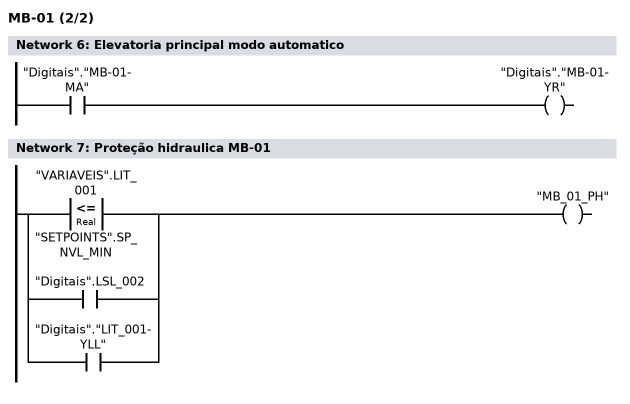
   RUNG wire#powerrail
      Contact( "Digitais"."MB-01-MA" )
      Coil( "Digitais"."MB-01-YR" )
   END_RUNG
   // the same network as SCL:
   "Digitais"."MB-01-YR" := "Digitais"."MB-01-MA";
END_REGION

REGION Network 7: Proteção hidraulica MB-01
   RUNG wire#powerrail
      { S7_Templates := "SrcType := Real" } LE_Contact(in1 := "VARIAVEIS".LIT_001, in2 := "SETPOINTS".SP_NVL_MIN)
      wire#w1
      Coil( "MB_01_PH" )
   END_RUNG
   RUNG wire#powerrail
      Contact( "Digitais".LSL_002 )
   END_RUNG wire#w1
   RUNG wire#powerrail
      Contact( "Digitais"."LIT_001-YLL" )
   END_RUNG wire#w1
   // the same network as SCL:
   "MB_01_PH" := ("VARIAVEIS".LIT_001 <= "SETPOINTS".SP_NVL_MIN) OR "Digitais".LSL_002 OR "Digitais"."LIT_001-YLL";
END_REGION
END_FUNCTION

FUNCTION "MB-02" : Void   // FC23, LAD
TITLE = Lógica de acionamento do motor
{ S7_Optimized_Access := 'FALSE' }
VERSION : 0.1
   VAR_TEMP
      IM : Bool;   // Intertravamento manual = 0
      IA : Bool;   // Intertravamento automáticol = 0
      HABM : Bool;   // Habilita funcionamento manual = 1
      HABA : Bool;   // Habilita funcionamento automático = 1
      CLM : Bool;   // Comando liga motor
      PROT : Bool;   // Proteção do motor acionada
   END_VAR
BEGIN

REGION Network 1: Intertravamento maual/automático
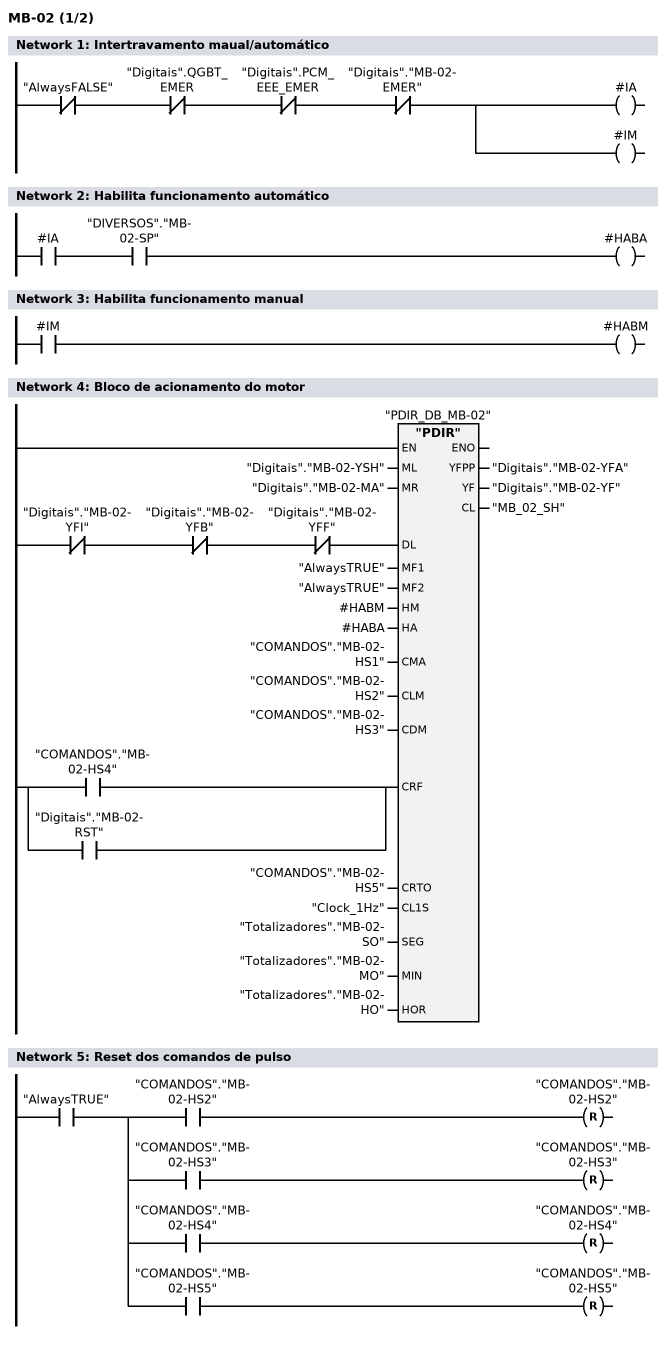
   RUNG wire#powerrail
      I_Contact( "AlwaysFALSE" )
      I_Contact( "Digitais".QGBT_EMER )
      I_Contact( "Digitais".PCM_EEE_EMER )
      I_Contact( "Digitais"."MB-02-EMER" )
      wire#w1
      Coil( #IA )
   END_RUNG
   RUNG wire#w1
      Coil( #IM )
   END_RUNG
   // the same network as SCL:
   #IA := NOT "AlwaysFALSE" AND NOT "Digitais".QGBT_EMER AND NOT "Digitais".PCM_EEE_EMER AND NOT "Digitais"."MB-02-EMER";
   #IM := #IA;
END_REGION

REGION Network 2: Habilita funcionamento automático
   RUNG wire#powerrail
      Contact( #IA )
      Contact( "DIVERSOS"."MB-02-SP" )
      Coil( #HABA )
   END_RUNG
   // the same network as SCL:
   #HABA := #IA AND "DIVERSOS"."MB-02-SP";
END_REGION

REGION Network 3: Habilita funcionamento manual
   RUNG wire#powerrail
      Contact( #IM )
      Coil( #HABM )
   END_RUNG
   // the same network as SCL:
   #HABM := #IM;
END_REGION

REGION Network 4: Bloco de acionamento do motor
   RUNG wire#powerrail
      "PDIR_DB_MB-02"(DL := wire#w1, CRF := wire#w2, ML := "Digitais"."MB-02-YSH", MR := "Digitais"."MB-02-MA", MF1 := "AlwaysTRUE", MF2 := "AlwaysTRUE", HM := #HABM, HA := #HABA, CMA := "COMANDOS"."MB-02-HS1", CLM := "COMANDOS"."MB-02-HS2", CDM := "COMANDOS"."MB-02-HS3", CRTO := "COMANDOS"."MB-02-HS5", CL1S := "Clock_1Hz", SEG := "Totalizadores"."MB-02-SO", MIN := "Totalizadores"."MB-02-MO", HOR := "Totalizadores"."MB-02-HO", YFPP => "Digitais"."MB-02-YFA", YF => "Digitais"."MB-02-YF", CL => "MB_02_SH")
   END_RUNG
   RUNG wire#powerrail
      I_Contact( "Digitais"."MB-02-YFI" )
      I_Contact( "Digitais"."MB-02-YFB" )
      I_Contact( "Digitais"."MB-02-YFF" )
   END_RUNG wire#w1
   RUNG wire#powerrail
      Contact( "COMANDOS"."MB-02-HS4" )
   END_RUNG wire#w2
   RUNG wire#powerrail
      Contact( "Digitais"."MB-02-RST" )
   END_RUNG wire#w2
   // the same network as SCL:
   "PDIR_DB_MB-02"(ML := "Digitais"."MB-02-YSH",   // "PDIR"
                   MR := "Digitais"."MB-02-MA",
                   DL := NOT "Digitais"."MB-02-YFI" AND NOT "Digitais"."MB-02-YFB" AND NOT "Digitais"."MB-02-YFF",
                   MF1 := "AlwaysTRUE",
                   MF2 := "AlwaysTRUE",
                   HM := #HABM,
                   HA := #HABA,
                   CMA := "COMANDOS"."MB-02-HS1",
                   CLM := "COMANDOS"."MB-02-HS2",
                   CDM := "COMANDOS"."MB-02-HS3",
                   CRF := "COMANDOS"."MB-02-HS4" OR "Digitais"."MB-02-RST",
                   CRTO := "COMANDOS"."MB-02-HS5",
                   CL1S := "Clock_1Hz",
                   SEG := "Totalizadores"."MB-02-SO",
                   MIN := "Totalizadores"."MB-02-MO",
                   HOR := "Totalizadores"."MB-02-HO",
                   YFPP => "Digitais"."MB-02-YFA",
                   YF => "Digitais"."MB-02-YF",
                   CL => "MB_02_SH");
END_REGION

REGION Network 5: Reset dos comandos de pulso
   RUNG wire#powerrail
      Contact( "AlwaysTRUE" )
      wire#w1
      Contact( "COMANDOS"."MB-02-HS2" )
      R_Coil( "COMANDOS"."MB-02-HS2" )
   END_RUNG
   RUNG wire#w1
      Contact( "COMANDOS"."MB-02-HS3" )
      R_Coil( "COMANDOS"."MB-02-HS3" )
   END_RUNG
   RUNG wire#w1
      Contact( "COMANDOS"."MB-02-HS4" )
      R_Coil( "COMANDOS"."MB-02-HS4" )
   END_RUNG
   RUNG wire#w1
      Contact( "COMANDOS"."MB-02-HS5" )
      R_Coil( "COMANDOS"."MB-02-HS5" )
   END_RUNG
   // the same network as SCL:
   IF "AlwaysTRUE" AND "COMANDOS"."MB-02-HS2" THEN "COMANDOS"."MB-02-HS2" := FALSE; END_IF;
   IF "AlwaysTRUE" AND "COMANDOS"."MB-02-HS3" THEN "COMANDOS"."MB-02-HS3" := FALSE; END_IF;
   IF "AlwaysTRUE" AND "COMANDOS"."MB-02-HS4" THEN "COMANDOS"."MB-02-HS4" := FALSE; END_IF;
   IF "AlwaysTRUE" AND "COMANDOS"."MB-02-HS5" THEN "COMANDOS"."MB-02-HS5" := FALSE; END_IF;
END_REGION

REGION Network 6: Elevatoria principal modo automatico
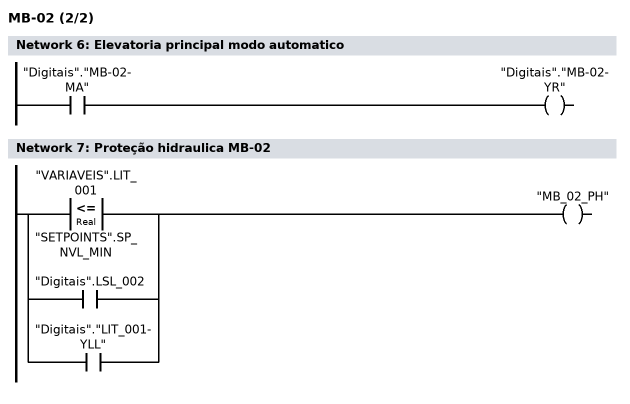
   RUNG wire#powerrail
      Contact( "Digitais"."MB-02-MA" )
      Coil( "Digitais"."MB-02-YR" )
   END_RUNG
   // the same network as SCL:
   "Digitais"."MB-02-YR" := "Digitais"."MB-02-MA";
END_REGION

REGION Network 7: Proteção hidraulica MB-02
   RUNG wire#powerrail
      { S7_Templates := "SrcType := Real" } LE_Contact(in1 := "VARIAVEIS".LIT_001, in2 := "SETPOINTS".SP_NVL_MIN)
      wire#w1
      Coil( "MB_02_PH" )
   END_RUNG
   RUNG wire#powerrail
      Contact( "Digitais".LSL_002 )
   END_RUNG wire#w1
   RUNG wire#powerrail
      Contact( "Digitais"."LIT_001-YLL" )
   END_RUNG wire#w1
   // the same network as SCL:
   "MB_02_PH" := ("VARIAVEIS".LIT_001 <= "SETPOINTS".SP_NVL_MIN) OR "Digitais".LSL_002 OR "Digitais"."LIT_001-YLL";
END_REGION
END_FUNCTION

FUNCTION "MB-03" : Void   // FC24, LAD
TITLE = Lógica de acionamento do motor
{ S7_Optimized_Access := 'FALSE' }
VERSION : 0.1
   VAR_TEMP
      IM : Bool;   // Intertravamento manual = 0
      IA : Bool;   // Intertravamento automáticol = 0
      HABM : Bool;   // Habilita funcionamento manual = 1
      HABA : Bool;   // Habilita funcionamento automático = 1
      CLM : Bool;   // Comando liga motor
      PROT : Bool;   // Proteção do motor acionada
   END_VAR
BEGIN

REGION Network 1: Intertravamento maual/automático
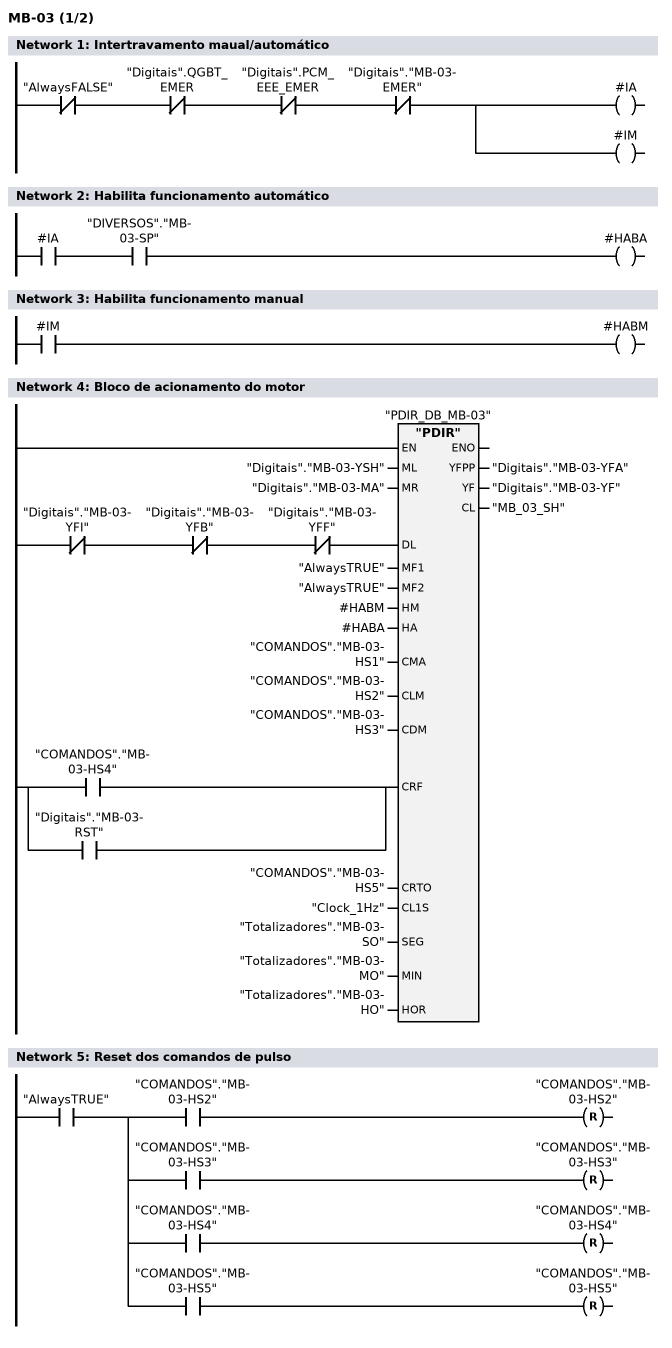
   RUNG wire#powerrail
      I_Contact( "AlwaysFALSE" )
      I_Contact( "Digitais".QGBT_EMER )
      I_Contact( "Digitais".PCM_EEE_EMER )
      I_Contact( "Digitais"."MB-03-EMER" )
      wire#w1
      Coil( #IA )
   END_RUNG
   RUNG wire#w1
      Coil( #IM )
   END_RUNG
   // the same network as SCL:
   #IA := NOT "AlwaysFALSE" AND NOT "Digitais".QGBT_EMER AND NOT "Digitais".PCM_EEE_EMER AND NOT "Digitais"."MB-03-EMER";
   #IM := #IA;
END_REGION

REGION Network 2: Habilita funcionamento automático
   RUNG wire#powerrail
      Contact( #IA )
      Contact( "DIVERSOS"."MB-03-SP" )
      Coil( #HABA )
   END_RUNG
   // the same network as SCL:
   #HABA := #IA AND "DIVERSOS"."MB-03-SP";
END_REGION

REGION Network 3: Habilita funcionamento manual
   RUNG wire#powerrail
      Contact( #IM )
      Coil( #HABM )
   END_RUNG
   // the same network as SCL:
   #HABM := #IM;
END_REGION

REGION Network 4: Bloco de acionamento do motor
   RUNG wire#powerrail
      "PDIR_DB_MB-03"(DL := wire#w1, CRF := wire#w2, ML := "Digitais"."MB-03-YSH", MR := "Digitais"."MB-03-MA", MF1 := "AlwaysTRUE", MF2 := "AlwaysTRUE", HM := #HABM, HA := #HABA, CMA := "COMANDOS"."MB-03-HS1", CLM := "COMANDOS"."MB-03-HS2", CDM := "COMANDOS"."MB-03-HS3", CRTO := "COMANDOS"."MB-03-HS5", CL1S := "Clock_1Hz", SEG := "Totalizadores"."MB-03-SO", MIN := "Totalizadores"."MB-03-MO", HOR := "Totalizadores"."MB-03-HO", YFPP => "Digitais"."MB-03-YFA", YF => "Digitais"."MB-03-YF", CL => "MB_03_SH")
   END_RUNG
   RUNG wire#powerrail
      I_Contact( "Digitais"."MB-03-YFI" )
      I_Contact( "Digitais"."MB-03-YFB" )
      I_Contact( "Digitais"."MB-03-YFF" )
   END_RUNG wire#w1
   RUNG wire#powerrail
      Contact( "COMANDOS"."MB-03-HS4" )
   END_RUNG wire#w2
   RUNG wire#powerrail
      Contact( "Digitais"."MB-03-RST" )
   END_RUNG wire#w2
   // the same network as SCL:
   "PDIR_DB_MB-03"(ML := "Digitais"."MB-03-YSH",   // "PDIR"
                   MR := "Digitais"."MB-03-MA",
                   DL := NOT "Digitais"."MB-03-YFI" AND NOT "Digitais"."MB-03-YFB" AND NOT "Digitais"."MB-03-YFF",
                   MF1 := "AlwaysTRUE",
                   MF2 := "AlwaysTRUE",
                   HM := #HABM,
                   HA := #HABA,
                   CMA := "COMANDOS"."MB-03-HS1",
                   CLM := "COMANDOS"."MB-03-HS2",
                   CDM := "COMANDOS"."MB-03-HS3",
                   CRF := "COMANDOS"."MB-03-HS4" OR "Digitais"."MB-03-RST",
                   CRTO := "COMANDOS"."MB-03-HS5",
                   CL1S := "Clock_1Hz",
                   SEG := "Totalizadores"."MB-03-SO",
                   MIN := "Totalizadores"."MB-03-MO",
                   HOR := "Totalizadores"."MB-03-HO",
                   YFPP => "Digitais"."MB-03-YFA",
                   YF => "Digitais"."MB-03-YF",
                   CL => "MB_03_SH");
END_REGION

REGION Network 5: Reset dos comandos de pulso
   RUNG wire#powerrail
      Contact( "AlwaysTRUE" )
      wire#w1
      Contact( "COMANDOS"."MB-03-HS2" )
      R_Coil( "COMANDOS"."MB-03-HS2" )
   END_RUNG
   RUNG wire#w1
      Contact( "COMANDOS"."MB-03-HS3" )
      R_Coil( "COMANDOS"."MB-03-HS3" )
   END_RUNG
   RUNG wire#w1
      Contact( "COMANDOS"."MB-03-HS4" )
      R_Coil( "COMANDOS"."MB-03-HS4" )
   END_RUNG
   RUNG wire#w1
      Contact( "COMANDOS"."MB-03-HS5" )
      R_Coil( "COMANDOS"."MB-03-HS5" )
   END_RUNG
   // the same network as SCL:
   IF "AlwaysTRUE" AND "COMANDOS"."MB-03-HS2" THEN "COMANDOS"."MB-03-HS2" := FALSE; END_IF;
   IF "AlwaysTRUE" AND "COMANDOS"."MB-03-HS3" THEN "COMANDOS"."MB-03-HS3" := FALSE; END_IF;
   IF "AlwaysTRUE" AND "COMANDOS"."MB-03-HS4" THEN "COMANDOS"."MB-03-HS4" := FALSE; END_IF;
   IF "AlwaysTRUE" AND "COMANDOS"."MB-03-HS5" THEN "COMANDOS"."MB-03-HS5" := FALSE; END_IF;
END_REGION

REGION Network 6: Elevatoria principal modo automatico
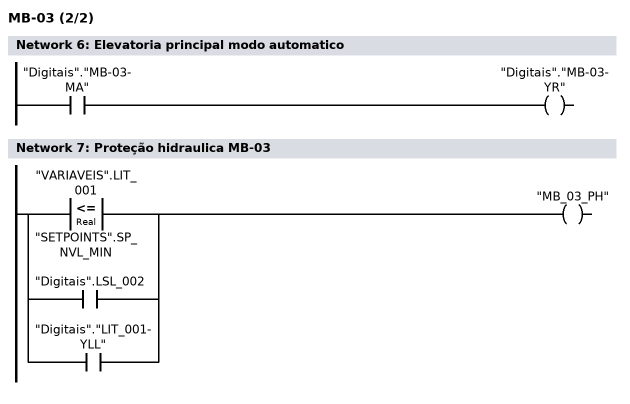
   RUNG wire#powerrail
      Contact( "Digitais"."MB-03-MA" )
      Coil( "Digitais"."MB-03-YR" )
   END_RUNG
   // the same network as SCL:
   "Digitais"."MB-03-YR" := "Digitais"."MB-03-MA";
END_REGION

REGION Network 7: Proteção hidraulica MB-03
   RUNG wire#powerrail
      { S7_Templates := "SrcType := Real" } LE_Contact(in1 := "VARIAVEIS".LIT_001, in2 := "SETPOINTS".SP_NVL_MIN)
      wire#w1
      Coil( "MB_03_PH" )
   END_RUNG
   RUNG wire#powerrail
      Contact( "Digitais".LSL_002 )
   END_RUNG wire#w1
   RUNG wire#powerrail
      Contact( "Digitais"."LIT_001-YLL" )
   END_RUNG wire#w1
   // the same network as SCL:
   "MB_03_PH" := ("VARIAVEIS".LIT_001 <= "SETPOINTS".SP_NVL_MIN) OR "Digitais".LSL_002 OR "Digitais"."LIT_001-YLL";
END_REGION
END_FUNCTION

FUNCTION "MB-04" : Void   // FC25, LAD
TITLE = Lógica de acionamento do motor
{ S7_Optimized_Access := 'FALSE' }
VERSION : 0.1
   VAR_TEMP
      IM : Bool;   // Intertravamento manual = 0
      IA : Bool;   // Intertravamento automáticol = 0
      HABM : Bool;   // Habilita funcionamento manual = 1
      HABA : Bool;   // Habilita funcionamento automático = 1
      CLM : Bool;   // Comando liga motor
      PROT : Bool;   // Proteção do motor acionada
   END_VAR
BEGIN

REGION Network 1: Intertravamento maual/automático
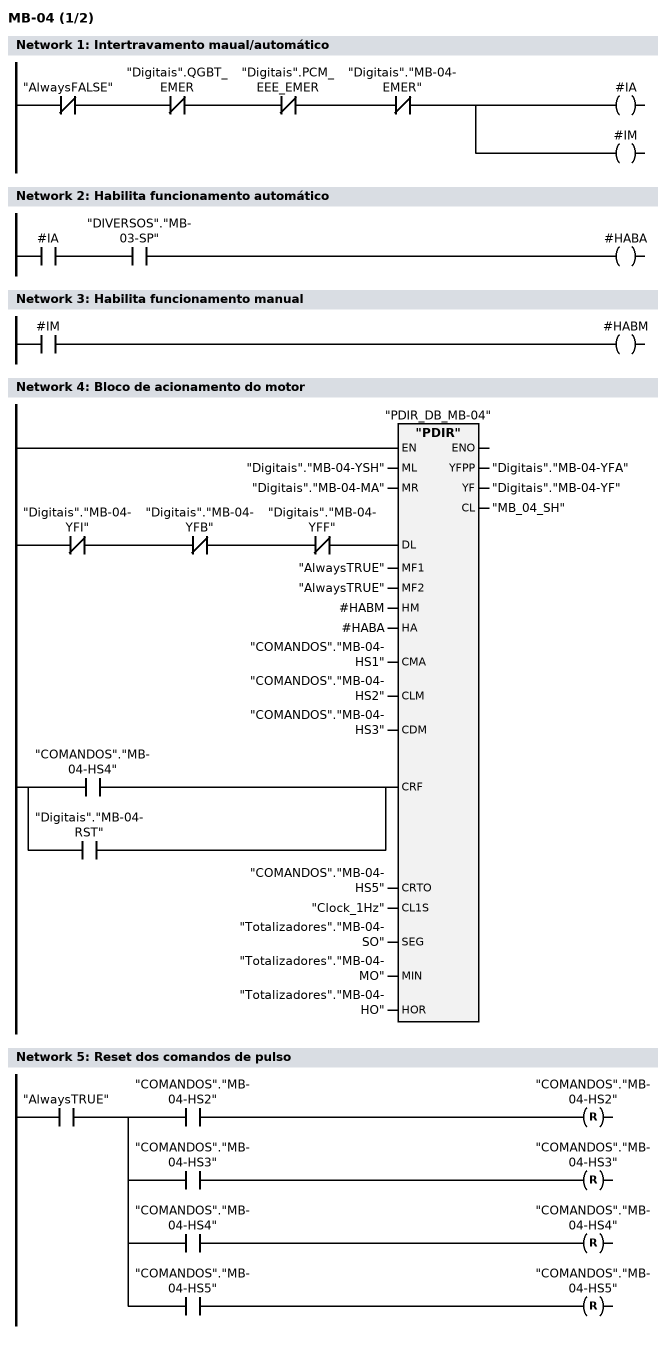
   RUNG wire#powerrail
      I_Contact( "AlwaysFALSE" )
      I_Contact( "Digitais".QGBT_EMER )
      I_Contact( "Digitais".PCM_EEE_EMER )
      I_Contact( "Digitais"."MB-04-EMER" )
      wire#w1
      Coil( #IA )
   END_RUNG
   RUNG wire#w1
      Coil( #IM )
   END_RUNG
   // the same network as SCL:
   #IA := NOT "AlwaysFALSE" AND NOT "Digitais".QGBT_EMER AND NOT "Digitais".PCM_EEE_EMER AND NOT "Digitais"."MB-04-EMER";
   #IM := #IA;
END_REGION

REGION Network 2: Habilita funcionamento automático
   RUNG wire#powerrail
      Contact( #IA )
      Contact( "DIVERSOS"."MB-03-SP" )
      Coil( #HABA )
   END_RUNG
   // the same network as SCL:
   #HABA := #IA AND "DIVERSOS"."MB-03-SP";
END_REGION

REGION Network 3: Habilita funcionamento manual
   RUNG wire#powerrail
      Contact( #IM )
      Coil( #HABM )
   END_RUNG
   // the same network as SCL:
   #HABM := #IM;
END_REGION

REGION Network 4: Bloco de acionamento do motor
   RUNG wire#powerrail
      "PDIR_DB_MB-04"(DL := wire#w1, CRF := wire#w2, ML := "Digitais"."MB-04-YSH", MR := "Digitais"."MB-04-MA", MF1 := "AlwaysTRUE", MF2 := "AlwaysTRUE", HM := #HABM, HA := #HABA, CMA := "COMANDOS"."MB-04-HS1", CLM := "COMANDOS"."MB-04-HS2", CDM := "COMANDOS"."MB-04-HS3", CRTO := "COMANDOS"."MB-04-HS5", CL1S := "Clock_1Hz", SEG := "Totalizadores"."MB-04-SO", MIN := "Totalizadores"."MB-04-MO", HOR := "Totalizadores"."MB-04-HO", YFPP => "Digitais"."MB-04-YFA", YF => "Digitais"."MB-04-YF", CL => "MB_04_SH")
   END_RUNG
   RUNG wire#powerrail
      I_Contact( "Digitais"."MB-04-YFI" )
      I_Contact( "Digitais"."MB-04-YFB" )
      I_Contact( "Digitais"."MB-04-YFF" )
   END_RUNG wire#w1
   RUNG wire#powerrail
      Contact( "COMANDOS"."MB-04-HS4" )
   END_RUNG wire#w2
   RUNG wire#powerrail
      Contact( "Digitais"."MB-04-RST" )
   END_RUNG wire#w2
   // the same network as SCL:
   "PDIR_DB_MB-04"(ML := "Digitais"."MB-04-YSH",   // "PDIR"
                   MR := "Digitais"."MB-04-MA",
                   DL := NOT "Digitais"."MB-04-YFI" AND NOT "Digitais"."MB-04-YFB" AND NOT "Digitais"."MB-04-YFF",
                   MF1 := "AlwaysTRUE",
                   MF2 := "AlwaysTRUE",
                   HM := #HABM,
                   HA := #HABA,
                   CMA := "COMANDOS"."MB-04-HS1",
                   CLM := "COMANDOS"."MB-04-HS2",
                   CDM := "COMANDOS"."MB-04-HS3",
                   CRF := "COMANDOS"."MB-04-HS4" OR "Digitais"."MB-04-RST",
                   CRTO := "COMANDOS"."MB-04-HS5",
                   CL1S := "Clock_1Hz",
                   SEG := "Totalizadores"."MB-04-SO",
                   MIN := "Totalizadores"."MB-04-MO",
                   HOR := "Totalizadores"."MB-04-HO",
                   YFPP => "Digitais"."MB-04-YFA",
                   YF => "Digitais"."MB-04-YF",
                   CL => "MB_04_SH");
END_REGION

REGION Network 5: Reset dos comandos de pulso
   RUNG wire#powerrail
      Contact( "AlwaysTRUE" )
      wire#w1
      Contact( "COMANDOS"."MB-04-HS2" )
      R_Coil( "COMANDOS"."MB-04-HS2" )
   END_RUNG
   RUNG wire#w1
      Contact( "COMANDOS"."MB-04-HS3" )
      R_Coil( "COMANDOS"."MB-04-HS3" )
   END_RUNG
   RUNG wire#w1
      Contact( "COMANDOS"."MB-04-HS4" )
      R_Coil( "COMANDOS"."MB-04-HS4" )
   END_RUNG
   RUNG wire#w1
      Contact( "COMANDOS"."MB-04-HS5" )
      R_Coil( "COMANDOS"."MB-04-HS5" )
   END_RUNG
   // the same network as SCL:
   IF "AlwaysTRUE" AND "COMANDOS"."MB-04-HS2" THEN "COMANDOS"."MB-04-HS2" := FALSE; END_IF;
   IF "AlwaysTRUE" AND "COMANDOS"."MB-04-HS3" THEN "COMANDOS"."MB-04-HS3" := FALSE; END_IF;
   IF "AlwaysTRUE" AND "COMANDOS"."MB-04-HS4" THEN "COMANDOS"."MB-04-HS4" := FALSE; END_IF;
   IF "AlwaysTRUE" AND "COMANDOS"."MB-04-HS5" THEN "COMANDOS"."MB-04-HS5" := FALSE; END_IF;
END_REGION

REGION Network 6: Elevatoria principal modo automatico
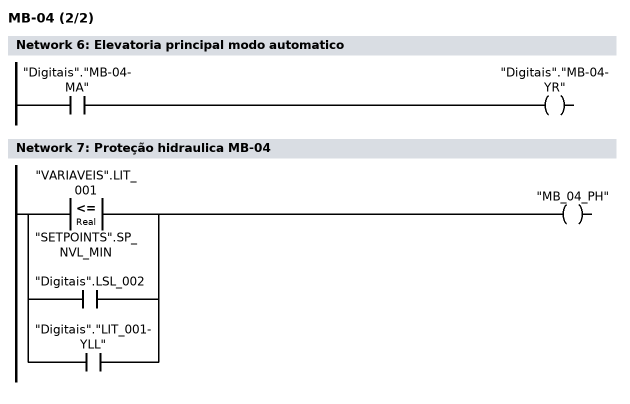
   RUNG wire#powerrail
      Contact( "Digitais"."MB-04-MA" )
      Coil( "Digitais"."MB-04-YR" )
   END_RUNG
   // the same network as SCL:
   "Digitais"."MB-04-YR" := "Digitais"."MB-04-MA";
END_REGION

REGION Network 7: Proteção hidraulica MB-04
   RUNG wire#powerrail
      { S7_Templates := "SrcType := Real" } LE_Contact(in1 := "VARIAVEIS".LIT_001, in2 := "SETPOINTS".SP_NVL_MIN)
      wire#w1
      Coil( "MB_04_PH" )
   END_RUNG
   RUNG wire#powerrail
      Contact( "Digitais".LSL_002 )
   END_RUNG wire#w1
   RUNG wire#powerrail
      Contact( "Digitais"."LIT_001-YLL" )
   END_RUNG wire#w1
   // the same network as SCL:
   "MB_04_PH" := ("VARIAVEIS".LIT_001 <= "SETPOINTS".SP_NVL_MIN) OR "Digitais".LSL_002 OR "Digitais"."LIT_001-YLL";
END_REGION
END_FUNCTION

ORGANIZATION_BLOCK "Main"   // OB1, LAD, ProgramCycle
TITLE = "Main Program Sweep (Cycle)"
{ S7_Optimized_Access := 'TRUE' }
VERSION : 0.1
   VAR_INPUT
      Initial_Call : Bool;   // Initial call of this OB
      Remanence : Bool;   // =True, if remanent data are available
   END_VAR
BEGIN

REGION Network 1: PULSO 1 SEGUNDO
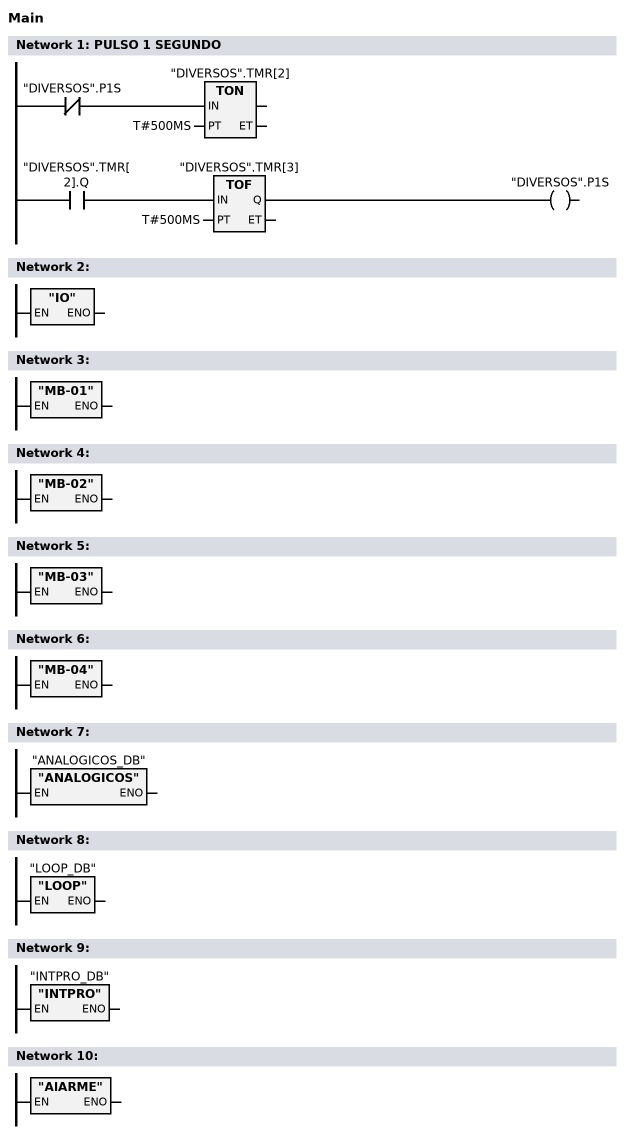
   "DIVERSOS".TMR[2].TON(IN := NOT "DIVERSOS".P1S, PT := T#500MS);
   "DIVERSOS".TMR[3].TOF(IN := "DIVERSOS".TMR[2].Q, PT := T#500MS);
   "DIVERSOS".P1S := "DIVERSOS".TMR[3].Q;
END_REGION

REGION Network 2
   RUNG wire#powerrail
      "IO"()
   END_RUNG
   // the same network as SCL:
   "IO"();
END_REGION

REGION Network 3
   RUNG wire#powerrail
      "MB-01"()
   END_RUNG
   // the same network as SCL:
   "MB-01"();
END_REGION

REGION Network 4
   RUNG wire#powerrail
      "MB-02"()
   END_RUNG
   // the same network as SCL:
   "MB-02"();
END_REGION

REGION Network 5
   RUNG wire#powerrail
      "MB-03"()
   END_RUNG
   // the same network as SCL:
   "MB-03"();
END_REGION

REGION Network 6
   RUNG wire#powerrail
      "MB-04"()
   END_RUNG
   // the same network as SCL:
   "MB-04"();
END_REGION

REGION Network 7
   RUNG wire#powerrail
      "ANALOGICOS_DB"()
   END_RUNG
   // the same network as SCL:
   "ANALOGICOS_DB"();   // "ANALOGICOS"
END_REGION

REGION Network 8
   RUNG wire#powerrail
      "LOOP_DB"()
   END_RUNG
   // the same network as SCL:
   "LOOP_DB"();   // "LOOP"
END_REGION

REGION Network 9
   RUNG wire#powerrail
      "INTPRO_DB"()
   END_RUNG
   // the same network as SCL:
   "INTPRO_DB"();   // "INTPRO"
END_REGION

REGION Network 10
   RUNG wire#powerrail
      "AlARME"()
   END_RUNG
   // the same network as SCL:
   "AlARME"();
END_REGION
END_ORGANIZATION_BLOCK

ORGANIZATION_BLOCK "CYC_INT5"   // OB35, LAD, CyclicInterrupt
TITLE = CONTROLE DE PID
{ S7_Optimized_Access := 'FALSE' }
VERSION : 0.1
   VAR_TEMP
      OB35_EV_CLASS : Byte;
      OB35_STRT_INF : Byte;
      OB35_PRIORITY : Byte;
      OB35_OB_NUMBR : Byte;
      OB35_RESERVED_1 : Byte;
      OB35_RESERVED_2 : Byte;
      OB35_PHASE_OFFSET : Word;
      OB35_RESERVED_3 : Int;
      OB35_EXC_FREQ : Int;
      OB35_DATE_TIME : Date_And_Time;
      "SPM-EEEB" : Real;   // Setpoint manual PID tanque de aeração 1
      EEEB_IT : Time;   // Ajuste integral do PID
      EEEB_DT : Time;   // Ajuste derivativo do PID
      EEEB_AUX : Real;   // Setpoint manual PID - auxiliar
      EEEB_P : Real;   // Setpoint manual PID - auxiliar
   END_VAR
   VAR_TEMP   // added for the SCL form of the ladder/FBD networks
      _w1 : Bool;
      _w2 : Bool;
      _w3 : Bool;
      _w4 : Bool;
   END_VAR
BEGIN

REGION Network 1 (STL): CONVERSÃO DOS SETPOINTS PARA TEMPO PID EEEB


   //CONVERSÃO DOS SETPOINTS DE TEMPO PID EEEB
         L     "PID"."PID-EEEB-I";
         L     1000.0;
         *R;
         RND;
         T     #EEEB_IT;

         L     "PID"."PID-EEEB-D";
         L     1000.0;
         *R;
         RND;
         T     #EEEB_DT;

         L     "PID"."PID-EEEB-P";
         L     -1.0;
         *R;
         T     #EEEB_P;
END_REGION

REGION Network 2: PID TANQUE DE AERAÇÃO 1
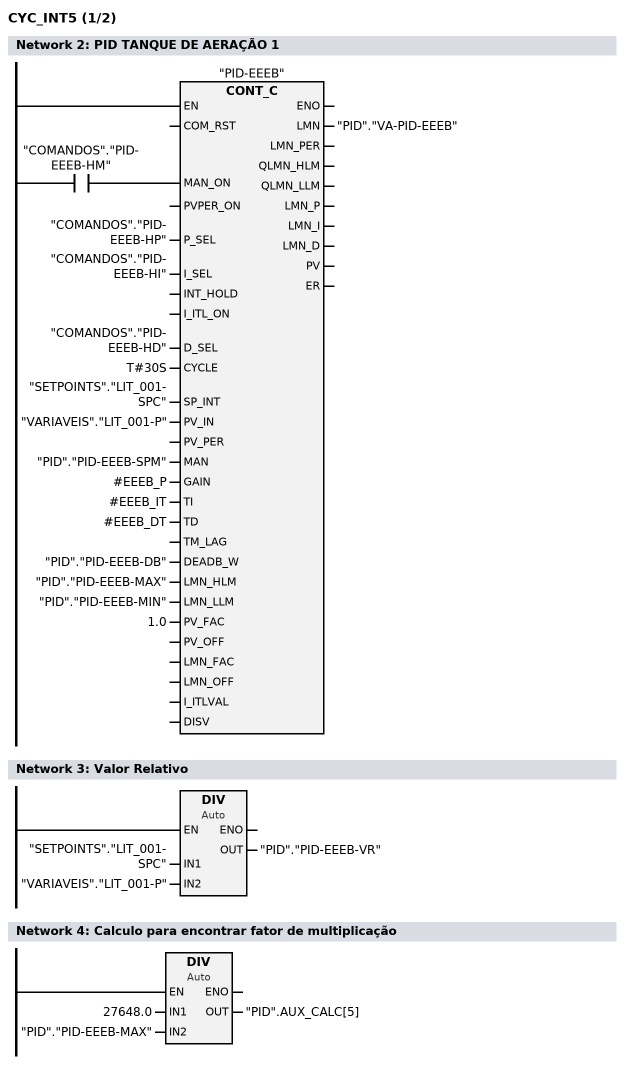
   "PID-EEEB"(MAN_ON := "COMANDOS"."PID-EEEB-HM",   // CONT_C
              P_SEL := "COMANDOS"."PID-EEEB-HP",
              I_SEL := "COMANDOS"."PID-EEEB-HI",
              D_SEL := "COMANDOS"."PID-EEEB-HD",
              CYCLE := T#30S,
              SP_INT := "SETPOINTS"."LIT_001-SPC",
              PV_IN := "VARIAVEIS"."LIT_001-P",
              MAN := "PID"."PID-EEEB-SPM",
              GAIN := #EEEB_P,
              TI := #EEEB_IT,
              TD := #EEEB_DT,
              DEADB_W := "PID"."PID-EEEB-DB",
              LMN_HLM := "PID"."PID-EEEB-MAX",
              LMN_LLM := "PID"."PID-EEEB-MIN",
              PV_FAC := 1.0,
              LMN => "PID"."VA-PID-EEEB");
END_REGION

REGION Network 3: Valor Relativo
   RUNG wire#powerrail
      Div(in1 := "SETPOINTS"."LIT_001-SPC", in2 := "VARIAVEIS"."LIT_001-P", out => "PID"."PID-EEEB-VR")
   END_RUNG
   // the same network as SCL:
   "PID"."PID-EEEB-VR" := "SETPOINTS"."LIT_001-SPC" / "VARIAVEIS"."LIT_001-P";
END_REGION

REGION Network 4: Calculo para encontrar fator de multiplicação
   RUNG wire#powerrail
      Div(in1 := 27648.0, in2 := "PID"."PID-EEEB-MAX", out => "PID".AUX_CALC[5])
   END_RUNG
   // the same network as SCL:
   "PID".AUX_CALC[5] := 27648.0 / "PID"."PID-EEEB-MAX";
END_REGION

REGION Network 5: Movimenta saida PID para entrada analógica inversor
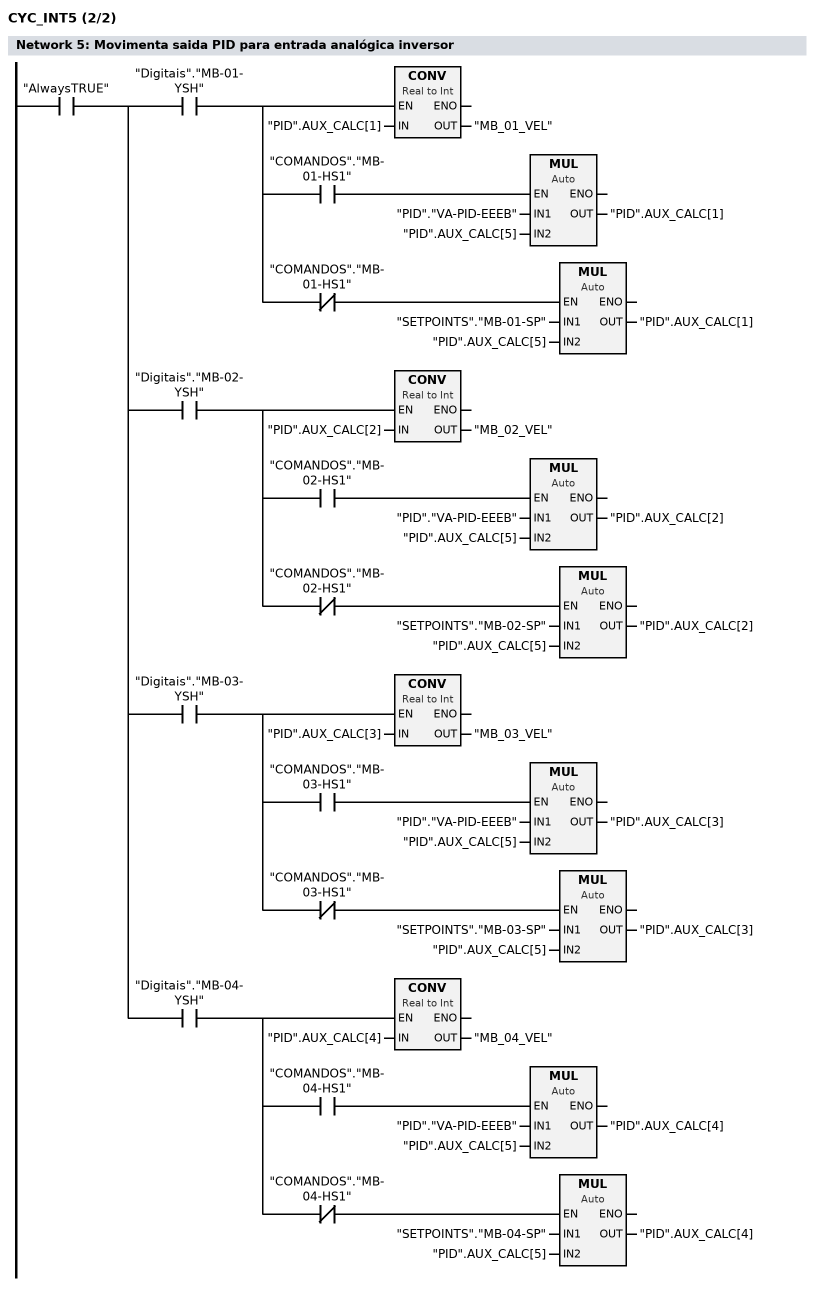
   RUNG wire#powerrail
      Contact( "AlwaysTRUE" )
      wire#w1
      Contact( "Digitais"."MB-01-YSH" )
      wire#w2
      { S7_Templates := "[SrcType := Real, DestType := Int]" } Convert(in := "PID".AUX_CALC[1], out => "MB_01_VEL")
   END_RUNG
   RUNG wire#w2
      Contact( "COMANDOS"."MB-01-HS1" )
      Mul(in1 := "PID"."VA-PID-EEEB", in2 := "PID".AUX_CALC[5], out => "PID".AUX_CALC[1])
   END_RUNG
   RUNG wire#w2
      I_Contact( "COMANDOS"."MB-01-HS1" )
      Mul(in1 := "SETPOINTS"."MB-01-SP", in2 := "PID".AUX_CALC[5], out => "PID".AUX_CALC[1])
   END_RUNG
   RUNG wire#w1
      Contact( "Digitais"."MB-02-YSH" )
      wire#w3
      { S7_Templates := "[SrcType := Real, DestType := Int]" } Convert(in := "PID".AUX_CALC[2], out => "MB_02_VEL")
   END_RUNG
   RUNG wire#w3
      Contact( "COMANDOS"."MB-02-HS1" )
      Mul(in1 := "PID"."VA-PID-EEEB", in2 := "PID".AUX_CALC[5], out => "PID".AUX_CALC[2])
   END_RUNG
   RUNG wire#w3
      I_Contact( "COMANDOS"."MB-02-HS1" )
      Mul(in1 := "SETPOINTS"."MB-02-SP", in2 := "PID".AUX_CALC[5], out => "PID".AUX_CALC[2])
   END_RUNG
   RUNG wire#w1
      Contact( "Digitais"."MB-03-YSH" )
      wire#w4
      { S7_Templates := "[SrcType := Real, DestType := Int]" } Convert(in := "PID".AUX_CALC[3], out => "MB_03_VEL")
   END_RUNG
   RUNG wire#w4
      Contact( "COMANDOS"."MB-03-HS1" )
      Mul(in1 := "PID"."VA-PID-EEEB", in2 := "PID".AUX_CALC[5], out => "PID".AUX_CALC[3])
   END_RUNG
   RUNG wire#w4
      I_Contact( "COMANDOS"."MB-03-HS1" )
      Mul(in1 := "SETPOINTS"."MB-03-SP", in2 := "PID".AUX_CALC[5], out => "PID".AUX_CALC[3])
   END_RUNG
   RUNG wire#w1
      Contact( "Digitais"."MB-04-YSH" )
      wire#w5
      { S7_Templates := "[SrcType := Real, DestType := Int]" } Convert(in := "PID".AUX_CALC[4], out => "MB_04_VEL")
   END_RUNG
   RUNG wire#w5
      Contact( "COMANDOS"."MB-04-HS1" )
      Mul(in1 := "PID"."VA-PID-EEEB", in2 := "PID".AUX_CALC[5], out => "PID".AUX_CALC[4])
   END_RUNG
   RUNG wire#w5
      I_Contact( "COMANDOS"."MB-04-HS1" )
      Mul(in1 := "SETPOINTS"."MB-04-SP", in2 := "PID".AUX_CALC[5], out => "PID".AUX_CALC[4])
   END_RUNG
   // the same network as SCL:
   #_w1 := "AlwaysTRUE" AND "Digitais"."MB-01-YSH";
   IF #_w1 THEN "MB_01_VEL" := REAL_TO_INT("PID".AUX_CALC[1]); END_IF;
   IF #_w1 AND "COMANDOS"."MB-01-HS1" THEN
       "PID".AUX_CALC[1] := "PID"."VA-PID-EEEB" * "PID".AUX_CALC[5];
   END_IF;
   IF #_w1 AND NOT "COMANDOS"."MB-01-HS1" THEN
       "PID".AUX_CALC[1] := "SETPOINTS"."MB-01-SP" * "PID".AUX_CALC[5];
   END_IF;
   #_w2 := "AlwaysTRUE" AND "Digitais"."MB-02-YSH";
   IF #_w2 THEN "MB_02_VEL" := REAL_TO_INT("PID".AUX_CALC[2]); END_IF;
   IF #_w2 AND "COMANDOS"."MB-02-HS1" THEN
       "PID".AUX_CALC[2] := "PID"."VA-PID-EEEB" * "PID".AUX_CALC[5];
   END_IF;
   IF #_w2 AND NOT "COMANDOS"."MB-02-HS1" THEN
       "PID".AUX_CALC[2] := "SETPOINTS"."MB-02-SP" * "PID".AUX_CALC[5];
   END_IF;
   #_w3 := "AlwaysTRUE" AND "Digitais"."MB-03-YSH";
   IF #_w3 THEN "MB_03_VEL" := REAL_TO_INT("PID".AUX_CALC[3]); END_IF;
   IF #_w3 AND "COMANDOS"."MB-03-HS1" THEN
       "PID".AUX_CALC[3] := "PID"."VA-PID-EEEB" * "PID".AUX_CALC[5];
   END_IF;
   IF #_w3 AND NOT "COMANDOS"."MB-03-HS1" THEN
       "PID".AUX_CALC[3] := "SETPOINTS"."MB-03-SP" * "PID".AUX_CALC[5];
   END_IF;
   #_w4 := "AlwaysTRUE" AND "Digitais"."MB-04-YSH";
   IF #_w4 THEN "MB_04_VEL" := REAL_TO_INT("PID".AUX_CALC[4]); END_IF;
   IF #_w4 AND "COMANDOS"."MB-04-HS1" THEN
       "PID".AUX_CALC[4] := "PID"."VA-PID-EEEB" * "PID".AUX_CALC[5];
   END_IF;
   IF #_w4 AND NOT "COMANDOS"."MB-04-HS1" THEN
       "PID".AUX_CALC[4] := "SETPOINTS"."MB-04-SP" * "PID".AUX_CALC[5];
   END_IF;
END_REGION
END_ORGANIZATION_BLOCK

(* ===== HMI "HMI_RT_1" =====
system functions are stored by id; their names below are inferred from use
connection "HMI_Connection_1": ETHERNET, SMART_S7_1500_OMS

HMI tags "Default tag table"
   "Digitais_MB-01-YSH" : Bool = PLC Digitais.MB-01-YSH AT %DB300.DBX0.0, 1 s
   "pause" : Bool = PLC pause AT %M2.1, 1 s
   "DIVERSOS_Looping" : Int = PLC DIVERSOS.Looping, 1 s
   "Tag_ScreenNumber" : Int, internal

HMI tags "ALARMES"
   "ALM0" : Word = PLC ALM0 AT %MW100, 1 s
   "ALM2" : Word = PLC ALM2 AT %MW102, 1 s
   "ALM4" : Word = PLC ALM4 AT %MW104, 1 s
   "ALM6" : Word = PLC ALM6 AT %MW106, 1 s
   "ALM8" : Word = PLC ALM8 AT %MW108, 1 s
   "ALM10" : Word = PLC ALM10 AT %MW110, 1 s
   "ALM12" : Word = PLC ALM12 AT %MW112, 1 s
   "ALM14" : Word = PLC ALM14 AT %MW114, 1 s
   "ALM16" : Word = PLC ALM16 AT %MW116, 1 s

HMI tags "PID"
   "PID_PID-EEEB-D" : Real = PLC PID.PID-EEEB-D AT %DB307.DBD0, 1 s
   "PID_PID-EEEB-P" : Real = PLC PID.PID-EEEB-P AT %DB307.DBD4, 1 s
   "PID_PID-EEEB-I" : Real = PLC PID.PID-EEEB-I AT %DB307.DBD8, 1 s
   "PID_PID-EEEB-MIN" : Real = PLC PID.PID-EEEB-MIN AT %DB307.DBD12, 1 s
   "PID_PID-EEEB-MAX" : Real = PLC PID.PID-EEEB-MAX AT %DB307.DBD16, 1 s
   "PID_PID-EEEB-DB" : Real = PLC PID.PID-EEEB-DB AT %DB307.DBD20, 1 s
   "PID_PID-EEEB-SPM" : Real = PLC PID.PID-EEEB-SPM AT %DB307.DBD24, 1 s
   "PID_VA-PID-EEEB" : Real = PLC PID.VA-PID-EEEB AT %DB307.DBD28, 1 s
   "PID_PID-EEEB-VR" : Real = PLC PID.PID-EEEB-VR AT %DB307.DBD32, 1 s

HMI tags "Comandos"
   "COMANDOS_MB-01-HS9" : Bool = PLC COMANDOS.MB-01-HS9 AT %DB303.DBX0.0, 1 s
   "COMANDOS_MB-01-HS10" : Bool = PLC COMANDOS.MB-01-HS10 AT %DB303.DBX0.1, 1 s
   "COMANDOS_MB-01-HS11" : Bool = PLC COMANDOS.MB-01-HS11 AT %DB303.DBX0.2, 1 s
   "COMANDOS_MB-01-HS12" : Bool = PLC COMANDOS.MB-01-HS12 AT %DB303.DBX0.3, 1 s
   "COMANDOS_MB-01-HS13" : Bool = PLC COMANDOS.MB-01-HS13 AT %DB303.DBX0.4, 1 s
   "COMANDOS_MB-01-HS14" : Bool = PLC COMANDOS.MB-01-HS14 AT %DB303.DBX0.5, 1 s
   "COMANDOS_MB-01-HS15" : Bool = PLC COMANDOS.MB-01-HS15 AT %DB303.DBX0.6, 1 s
   "COMANDOS_MB-01-HS16" : Bool = PLC COMANDOS.MB-01-HS16 AT %DB303.DBX0.7, 1 s
   "COMANDOS_MB-01-HS1" : Bool = PLC COMANDOS.MB-01-HS1 AT %DB303.DBX1.0, 1 s
   "COMANDOS_MB-01-HS2" : Bool = PLC COMANDOS.MB-01-HS2 AT %DB303.DBX1.1, 1 s
   "COMANDOS_MB-01-HS3" : Bool = PLC COMANDOS.MB-01-HS3 AT %DB303.DBX1.2, 1 s
   "COMANDOS_MB-01-HS4" : Bool = PLC COMANDOS.MB-01-HS4 AT %DB303.DBX1.3, 1 s
   "COMANDOS_MB-01-HS5" : Bool = PLC COMANDOS.MB-01-HS5 AT %DB303.DBX1.4, 1 s
   "COMANDOS_MB-01-HS6" : Bool = PLC COMANDOS.MB-01-HS6 AT %DB303.DBX1.5, 1 s
   "COMANDOS_MB-01-HS7" : Bool = PLC COMANDOS.MB-01-HS7 AT %DB303.DBX1.6, 1 s
   "COMANDOS_MB-01-HS8" : Bool = PLC COMANDOS.MB-01-HS8 AT %DB303.DBX1.7, 1 s
   "COMANDOS_MB-02-HS9" : Bool = PLC COMANDOS.MB-02-HS9 AT %DB303.DBX2.0, 1 s
   "COMANDOS_MB-02-HS10" : Bool = PLC COMANDOS.MB-02-HS10 AT %DB303.DBX2.1, 1 s
   "COMANDOS_MB-02-HS11" : Bool = PLC COMANDOS.MB-02-HS11 AT %DB303.DBX2.2, 1 s
   "COMANDOS_MB-02-HS12" : Bool = PLC COMANDOS.MB-02-HS12 AT %DB303.DBX2.3, 1 s
   "COMANDOS_MB-02-HS13" : Bool = PLC COMANDOS.MB-02-HS13 AT %DB303.DBX2.4, 1 s
   "COMANDOS_MB-02-HS14" : Bool = PLC COMANDOS.MB-02-HS14 AT %DB303.DBX2.5, 1 s
   "COMANDOS_MB-02-HS15" : Bool = PLC COMANDOS.MB-02-HS15 AT %DB303.DBX2.6, 1 s
   "COMANDOS_MB-02-HS16" : Bool = PLC COMANDOS.MB-02-HS16 AT %DB303.DBX2.7, 1 s
   "COMANDOS_MB-02-HS1" : Bool = PLC COMANDOS.MB-02-HS1 AT %DB303.DBX3.0, 1 s
   "COMANDOS_MB-02-HS2" : Bool = PLC COMANDOS.MB-02-HS2 AT %DB303.DBX3.1, 1 s
   "COMANDOS_MB-02-HS3" : Bool = PLC COMANDOS.MB-02-HS3 AT %DB303.DBX3.2, 1 s
   "COMANDOS_MB-02-HS4" : Bool = PLC COMANDOS.MB-02-HS4 AT %DB303.DBX3.3, 1 s
   "COMANDOS_MB-02-HS5" : Bool = PLC COMANDOS.MB-02-HS5 AT %DB303.DBX3.4, 1 s
   "COMANDOS_MB-02-HS6" : Bool = PLC COMANDOS.MB-02-HS6 AT %DB303.DBX3.5, 1 s
   "COMANDOS_MB-02-HS7" : Bool = PLC COMANDOS.MB-02-HS7 AT %DB303.DBX3.6, 1 s
   "COMANDOS_MB-02-HS8" : Bool = PLC COMANDOS.MB-02-HS8 AT %DB303.DBX3.7, 1 s
   "COMANDOS_MB-03-HS9" : Bool = PLC COMANDOS.MB-03-HS9 AT %DB303.DBX4.0, 1 s
   "COMANDOS_MB-03-HS10" : Bool = PLC COMANDOS.MB-03-HS10 AT %DB303.DBX4.1, 1 s
   "COMANDOS_MB-03-HS11" : Bool = PLC COMANDOS.MB-03-HS11 AT %DB303.DBX4.2, 1 s
   "COMANDOS_MB-03-HS12" : Bool = PLC COMANDOS.MB-03-HS12 AT %DB303.DBX4.3, 1 s
   "COMANDOS_MB-03-HS13" : Bool = PLC COMANDOS.MB-03-HS13 AT %DB303.DBX4.4, 1 s
   "COMANDOS_MB-03-HS14" : Bool = PLC COMANDOS.MB-03-HS14 AT %DB303.DBX4.5, 1 s
   "COMANDOS_MB-03-HS15" : Bool = PLC COMANDOS.MB-03-HS15 AT %DB303.DBX4.6, 1 s
   "COMANDOS_MB-03-HS16" : Bool = PLC COMANDOS.MB-03-HS16 AT %DB303.DBX4.7, 1 s
   "COMANDOS_MB-03-HS1" : Bool = PLC COMANDOS.MB-03-HS1 AT %DB303.DBX5.0, 1 s
   "COMANDOS_MB-03-HS2" : Bool = PLC COMANDOS.MB-03-HS2 AT %DB303.DBX5.1, 1 s
   "COMANDOS_MB-03-HS3" : Bool = PLC COMANDOS.MB-03-HS3 AT %DB303.DBX5.2, 1 s
   "COMANDOS_MB-03-HS4" : Bool = PLC COMANDOS.MB-03-HS4 AT %DB303.DBX5.3, 1 s
   "COMANDOS_MB-03-HS5" : Bool = PLC COMANDOS.MB-03-HS5 AT %DB303.DBX5.4, 1 s
   "COMANDOS_MB-03-HS6" : Bool = PLC COMANDOS.MB-03-HS6 AT %DB303.DBX5.5, 1 s
   "COMANDOS_MB-03-HS7" : Bool = PLC COMANDOS.MB-03-HS7 AT %DB303.DBX5.6, 1 s
   "COMANDOS_MB-03-HS8" : Bool = PLC COMANDOS.MB-03-HS8 AT %DB303.DBX5.7, 1 s
   "COMANDOS_MB-04-HS9" : Bool = PLC COMANDOS.MB-04-HS9 AT %DB303.DBX6.0, 1 s
   "COMANDOS_MB-04-HS10" : Bool = PLC COMANDOS.MB-04-HS10 AT %DB303.DBX6.1, 1 s
   "COMANDOS_MB-04-HS11" : Bool = PLC COMANDOS.MB-04-HS11 AT %DB303.DBX6.2, 1 s
   "COMANDOS_MB-04-HS12" : Bool = PLC COMANDOS.MB-04-HS12 AT %DB303.DBX6.3, 1 s
   "COMANDOS_MB-04-HS13" : Bool = PLC COMANDOS.MB-04-HS13 AT %DB303.DBX6.4, 1 s
   "COMANDOS_MB-04-HS14" : Bool = PLC COMANDOS.MB-04-HS14 AT %DB303.DBX6.5, 1 s
   "COMANDOS_MB-04-HS15" : Bool = PLC COMANDOS.MB-04-HS15 AT %DB303.DBX6.6, 1 s
   "COMANDOS_MB-04-HS16" : Bool = PLC COMANDOS.MB-04-HS16 AT %DB303.DBX6.7, 1 s
   "COMANDOS_MB-04-HS1" : Bool = PLC COMANDOS.MB-04-HS1 AT %DB303.DBX7.0, 1 s
   "COMANDOS_MB-04-HS2" : Bool = PLC COMANDOS.MB-04-HS2 AT %DB303.DBX7.1, 1 s
   "COMANDOS_MB-04-HS3" : Bool = PLC COMANDOS.MB-04-HS3 AT %DB303.DBX7.2, 1 s
   "COMANDOS_MB-04-HS4" : Bool = PLC COMANDOS.MB-04-HS4 AT %DB303.DBX7.3, 1 s
   "COMANDOS_MB-04-HS5" : Bool = PLC COMANDOS.MB-04-HS5 AT %DB303.DBX7.4, 1 s
   "COMANDOS_MB-04-HS6" : Bool = PLC COMANDOS.MB-04-HS6 AT %DB303.DBX7.5, 1 s
   "COMANDOS_MB-04-HS7" : Bool = PLC COMANDOS.MB-04-HS7 AT %DB303.DBX7.6, 1 s
   "COMANDOS_MB-04-HS8" : Bool = PLC COMANDOS.MB-04-HS8 AT %DB303.DBX7.7, 1 s
   "COMANDOS_LIT_001-HS9" : Bool = PLC COMANDOS.LIT_001-HS9 AT %DB303.DBX8.0, 1 s
   "COMANDOS_LIT_001-HS10" : Bool = PLC COMANDOS.LIT_001-HS10 AT %DB303.DBX8.1, 1 s
   "COMANDOS_LIT_001-HS11" : Bool = PLC COMANDOS.LIT_001-HS11 AT %DB303.DBX8.2, 1 s
   "COMANDOS_LIT_001-HS12" : Bool = PLC COMANDOS.LIT_001-HS12 AT %DB303.DBX8.3, 1 s
   "COMANDOS_LIT_001-HS13" : Bool = PLC COMANDOS.LIT_001-HS13 AT %DB303.DBX8.4, 1 s
   "COMANDOS_LIT_001-HS14" : Bool = PLC COMANDOS.LIT_001-HS14 AT %DB303.DBX8.5, 1 s
   "COMANDOS_LIT_001-HS15" : Bool = PLC COMANDOS.LIT_001-HS15 AT %DB303.DBX8.6, 1 s
   "COMANDOS_LIT_001-HS16" : Bool = PLC COMANDOS.LIT_001-HS16 AT %DB303.DBX8.7, 1 s
   "COMANDOS_LIT_001-HSHH" : Bool = PLC COMANDOS.LIT_001-HSHH AT %DB303.DBX9.0, 1 s
   "COMANDOS_LIT_001-HSH" : Bool = PLC COMANDOS.LIT_001-HSH AT %DB303.DBX9.1, 1 s
   "COMANDOS_LIT_001-HSL" : Bool = PLC COMANDOS.LIT_001-HSL AT %DB303.DBX9.2, 1 s
   "COMANDOS_LIT_001-HSLL" : Bool = PLC COMANDOS.LIT_001-HSLL AT %DB303.DBX9.3, 1 s
   "COMANDOS_LIT_001-HSM" : Bool = PLC COMANDOS.LIT_001-HSM AT %DB303.DBX9.4, 1 s
   "COMANDOS_LIT_001-HS6" : Bool = PLC COMANDOS.LIT_001-HS6 AT %DB303.DBX9.5, 1 s
   "COMANDOS_LIT_001-HS7" : Bool = PLC COMANDOS.LIT_001-HS7 AT %DB303.DBX9.6, 1 s
   "COMANDOS_LIT_001-HS8" : Bool = PLC COMANDOS.LIT_001-HS8 AT %DB303.DBX9.7, 1 s
   "COMANDOS_PID-EEEB-HD" : Bool = PLC COMANDOS.PID-EEEB-HD AT %DB303.DBX10.1, 1 s
   "COMANDOS_PID-EEEB-HP" : Bool = PLC COMANDOS.PID-EEEB-HP AT %DB303.DBX10.2, 1 s
   "COMANDOS_PID-EEEB-HI" : Bool = PLC COMANDOS.PID-EEEB-HI AT %DB303.DBX10.3, 1 s
   "COMANDOS_PID-EEEB-HM" : Bool = PLC COMANDOS.PID-EEEB-HM AT %DB303.DBX12.2, 1 s
